      Appearance <- "PN_PB\PTMUX_F_TLN113_128"
   TextField "OBJECT_484" at 1009,421 size 40x20; Text '115'
      Appearance <- "PN_PB\PTMUX_F_TLN113_128"
   GraphicIOField "OBJECT_485" at 936,410 size 60x43; PictureList "PB_Slave_Bit12_2"
      ProcessValue <- "PN_PB\PTMUX_P_TLN113_128"
   TextField "OBJECT_486" at 946,421 size 40x20; Text '116'
      Appearance <- "PN_PB\PTMUX_F_TLN113_128"
   GraphicIOField "OBJECT_488" at 748,410 size 60x43; PictureList "PB_Slave_Bit15_2"
      ProcessValue <- "PN_PB\PTMUX_P_TLN113_128"
   TextField "OBJECT_489" at 758,421 size 40x20; Text '119'
      Appearance <- "PN_PB\PTMUX_F_TLN113_128"
   GraphicIOField "OBJECT_210" at 246,89 size 60x43; PictureList "PB_Slave_Bit7_2"
      ProcessValue <- "PN_PB\PTMUX_P_TLN1_16"
   GraphicIOField "OBJECT_214" at 372,89 size 60x43; PictureList "PB_Slave_Bit5_2"
      ProcessValue <- "PN_PB\PTMUX_P_TLN1_16"
   GraphicIOField "OBJECT_215" at 434,89 size 60x43; PictureList "PB_Slave_Bit4_2"
      ProcessValue <- "PN_PB\PTMUX_P_TLN1_16"
   TextField "OBJECT_218" at 506,100 size 40x20; Text '1'
   GraphicIOField "OBJECT_219" at 560,89 size 60x43; PictureList "PB_Slave_Bit2_2"
      ProcessValue <- "PN_PB\PTMUX_P_TLN1_16"
   GraphicIOField "OBJECT_221" at 622,89 size 60x43; PictureList "PB_Slave_Bit1_2"
      ProcessValue <- "PN_PB\PTMUX_P_TLN1_16"
   GraphicIOField "OBJECT_222" at 685,89 size 60x43; PictureList "PB_Slave_Bit0_2"
      ProcessValue <- "PN_PB\PTMUX_P_TLN1_16"
   TextField "OBJECT_223" at 696,100 size 40x20; Text '8'
      Appearance <- "PN_PB\PTMUX_F_TLN1_16"
   GraphicIOField "OBJECT_225" at 497,89 size 60x43; PictureList "PB_Slave_Bit3_2"
      ProcessValue <- "PN_PB\PTMUX_P_TLN1_16"
   TextField "OBJECT_226" at 633,100 size 40x20; Text '9'
      Appearance <- "PN_PB\PTMUX_F_TLN1_16"
   TextField "OBJECT_227" at 570,100 size 40x20; Text '10'
      Appearance <- "PN_PB\PTMUX_F_TLN1_16"
   TextField "OBJECT_228" at 508,100 size 40x20; Text '11'
      Appearance <- "PN_PB\PTMUX_F_TLN1_16"
   TextField "OBJECT_229" at 445,100 size 40x20; Text '12'
      Appearance <- "PN_PB\PTMUX_F_TLN1_16"
   TextField "OBJECT_230" at 382,100 size 40x20; Text '13'
      Appearance <- "PN_PB\PTMUX_F_TLN1_16"
   TextField "OBJECT_231" at 320,100 size 40x20; Text '14'
      Appearance <- "PN_PB\PTMUX_F_TLN1_16"
   TextField "OBJECT_232" at 257,100 size 40x20; Text '15'
      Appearance <- "PN_PB\PTMUX_F_TLN1_16"
   GraphicIOField "OBJECT_250" at 246,134 size 60x43; PictureList "PB_Slave_Bit7_2"
      ProcessValue <- "PN_PB\PTMUX_P_TLN17_32"
   GraphicIOField "OBJECT_251" at 309,134 size 60x43; PictureList "PB_Slave_Bit6_2"
      ProcessValue <- "PN_PB\PTMUX_P_TLN17_32"
   GraphicIOField "OBJECT_252" at 372,134 size 60x43; PictureList "PB_Slave_Bit5_2"
      ProcessValue <- "PN_PB\PTMUX_P_TLN17_32"
   GraphicIOField "OBJECT_253" at 434,134 size 60x43; PictureList "PB_Slave_Bit4_2"
      ProcessValue <- "PN_PB\PTMUX_P_TLN17_32"
   TextField "OBJECT_254" at 506,145 size 40x20; Text '1'
   GraphicIOField "OBJECT_255" at 560,134 size 60x43; PictureList "PB_Slave_Bit2_2"
      ProcessValue <- "PN_PB\PTMUX_P_TLN17_32"
   GraphicIOField "OBJECT_256" at 622,134 size 60x43; PictureList "PB_Slave_Bit1_2"
      ProcessValue <- "PN_PB\PTMUX_P_TLN17_32"
   GraphicIOField "OBJECT_257" at 685,134 size 60x43; PictureList "PB_Slave_Bit0_2"
      ProcessValue <- "PN_PB\PTMUX_P_TLN17_32"
   TextField "OBJECT_258" at 696,145 size 40x20; Text '24'
      Appearance <- "PN_PB\PTMUX_F_TLN17_32"
   GraphicIOField "OBJECT_259" at 497,134 size 60x43; PictureList "PB_Slave_Bit3_2"
      ProcessValue <- "PN_PB\PTMUX_P_TLN17_32"
   TextField "OBJECT_260" at 633,145 size 40x20; Text '25'
      Appearance <- "PN_PB\PTMUX_F_TLN17_32"
   TextField "OBJECT_261" at 570,145 size 40x20; Text '26'
      Appearance <- "PN_PB\PTMUX_F_TLN17_32"
   TextField "OBJECT_262" at 508,145 size 40x20; Text '27'
      Appearance <- "PN_PB\PTMUX_F_TLN17_32"
   TextField "OBJECT_263" at 445,145 size 40x20; Text '28'
      Appearance <- "PN_PB\PTMUX_F_TLN17_32"
   TextField "OBJECT_264" at 382,145 size 40x20; Text '29'
      Appearance <- "PN_PB\PTMUX_F_TLN17_32"
   TextField "OBJECT_265" at 320,145 size 40x20; Text '30'
      Appearance <- "PN_PB\PTMUX_F_TLN17_32"
   TextField "OBJECT_266" at 257,145 size 40x20; Text '31'
      Appearance <- "PN_PB\PTMUX_F_TLN17_32"
   GraphicIOField "OBJECT_283" at 246,180 size 60x43; PictureList "PB_Slave_Bit7_2"
      ProcessValue <- "PN_PB\PTMUX_P_TLN33_48"
   GraphicIOField "OBJECT_284" at 309,180 size 60x43; PictureList "PB_Slave_Bit6_2"
      ProcessValue <- "PN_PB\PTMUX_P_TLN33_48"
   GraphicIOField "OBJECT_285" at 372,180 size 60x43; PictureList "PB_Slave_Bit5_2"
      ProcessValue <- "PN_PB\PTMUX_P_TLN33_48"
   GraphicIOField "OBJECT_286" at 434,180 size 60x43; PictureList "PB_Slave_Bit4_2"
      ProcessValue <- "PN_PB\PTMUX_P_TLN33_48"
   TextField "OBJECT_287" at 506,190 size 40x20; Text '1'
   GraphicIOField "OBJECT_288" at 560,180 size 60x43; PictureList "PB_Slave_Bit2_2"
      ProcessValue <- "PN_PB\PTMUX_P_TLN33_48"
   GraphicIOField "OBJECT_289" at 622,180 size 60x43; PictureList "PB_Slave_Bit1_2"
      ProcessValue <- "PN_PB\PTMUX_P_TLN33_48"
   GraphicIOField "OBJECT_290" at 685,180 size 60x43; PictureList "PB_Slave_Bit0_2"
      ProcessValue <- "PN_PB\PTMUX_P_TLN33_48"
   TextField "OBJECT_291" at 696,190 size 40x20; Text '40'
      Appearance <- "PN_PB\PTMUX_F_TLN33_48"
   GraphicIOField "OBJECT_292" at 497,180 size 60x43; PictureList "PB_Slave_Bit3_2"
      ProcessValue <- "PN_PB\PTMUX_P_TLN33_48"
   TextField "OBJECT_293" at 633,190 size 40x20; Text '41'
      Appearance <- "PN_PB\PTMUX_F_TLN33_48"
   TextField "OBJECT_294" at 570,190 size 40x20; Text '42'
      Appearance <- "PN_PB\PTMUX_F_TLN33_48"
   TextField "OBJECT_295" at 508,190 size 40x20; Text '43'
      Appearance <- "PN_PB\PTMUX_F_TLN33_48"
   TextField "OBJECT_296" at 445,190 size 40x20; Text '44'
      Appearance <- "PN_PB\PTMUX_F_TLN33_48"
   TextField "OBJECT_297" at 382,190 size 40x20; Text '45'
      Appearance <- "PN_PB\PTMUX_F_TLN33_48"
   TextField "OBJECT_298" at 320,190 size 40x20; Text '46'
      Appearance <- "PN_PB\PTMUX_F_TLN33_48"
   TextField "OBJECT_299" at 257,190 size 40x20; Text '47'
      Appearance <- "PN_PB\PTMUX_F_TLN33_48"
   GraphicIOField "OBJECT_318" at 246,225 size 60x43; PictureList "PB_Slave_Bit7_2"
      ProcessValue <- "PN_PB\PTMUX_P_TLN49_64"
   GraphicIOField "OBJECT_319" at 309,225 size 60x43; PictureList "PB_Slave_Bit6_2"
      ProcessValue <- "PN_PB\PTMUX_P_TLN49_64"
   GraphicIOField "OBJECT_320" at 372,225 size 60x43; PictureList "PB_Slave_Bit5_2"
      ProcessValue <- "PN_PB\PTMUX_P_TLN49_64"
   GraphicIOField "OBJECT_321" at 434,225 size 60x43; PictureList "PB_Slave_Bit4_2"
      ProcessValue <- "PN_PB\PTMUX_P_TLN49_64"
   TextField "OBJECT_322" at 506,236 size 40x20; Text '1'
   GraphicIOField "OBJECT_323" at 560,225 size 60x43; PictureList "PB_Slave_Bit2_2"
      ProcessValue <- "PN_PB\PTMUX_P_TLN49_64"
   GraphicIOField "OBJECT_324" at 622,225 size 60x43; PictureList "PB_Slave_Bit1_2"
      ProcessValue <- "PN_PB\PTMUX_P_TLN49_64"
   GraphicIOField "OBJECT_325" at 685,225 size 60x43; PictureList "PB_Slave_Bit0_2"
      ProcessValue <- "PN_PB\PTMUX_P_TLN49_64"
   TextField "OBJECT_326" at 696,236 size 40x20; Text '56'
      Appearance <- "PN_PB\PTMUX_F_TLN49_64"
   GraphicIOField "OBJECT_327" at 497,225 size 60x43; PictureList "PB_Slave_Bit3_2"
      ProcessValue <- "PN_PB\PTMUX_P_TLN49_64"
   TextField "OBJECT_328" at 633,236 size 40x20; Text '57'
      Appearance <- "PN_PB\PTMUX_F_TLN49_64"
   TextField "OBJECT_329" at 570,236 size 40x20; Text '58'
      Appearance <- "PN_PB\PTMUX_F_TLN49_64"
   TextField "OBJECT_330" at 508,236 size 40x20; Text '59'
      Appearance <- "PN_PB\PTMUX_F_TLN49_64"
   TextField "OBJECT_331" at 445,236 size 40x20; Text '60'
      Appearance <- "PN_PB\PTMUX_F_TLN49_64"
   TextField "OBJECT_332" at 382,236 size 40x20; Text '61'
      Appearance <- "PN_PB\PTMUX_F_TLN49_64"
   TextField "OBJECT_333" at 320,236 size 40x20; Text '62'
      Appearance <- "PN_PB\PTMUX_F_TLN49_64"
   TextField "OBJECT_334" at 257,236 size 40x20; Text '63'
      Appearance <- "PN_PB\PTMUX_F_TLN49_64"
   GraphicIOField "OBJECT_352" at 246,270 size 60x43; PictureList "PB_Slave_Bit7_2"
      ProcessValue <- "PN_PB\PTMUX_P_TLN65_80"
   GraphicIOField "OBJECT_353" at 309,270 size 60x43; PictureList "PB_Slave_Bit6_2"
      ProcessValue <- "PN_PB\PTMUX_P_TLN65_80"
   GraphicIOField "OBJECT_354" at 372,270 size 60x43; PictureList "PB_Slave_Bit5_2"
      ProcessValue <- "PN_PB\PTMUX_P_TLN65_80"
   GraphicIOField "OBJECT_355" at 434,270 size 60x43; PictureList "PB_Slave_Bit4_2"
      ProcessValue <- "PN_PB\PTMUX_P_TLN65_80"
   TextField "OBJECT_356" at 506,282 size 40x20; Text '1'
   GraphicIOField "OBJECT_357" at 560,270 size 60x43; PictureList "PB_Slave_Bit2_2"
      ProcessValue <- "PN_PB\PTMUX_P_TLN65_80"
   GraphicIOField "OBJECT_358" at 622,270 size 60x43; PictureList "PB_Slave_Bit1_2"
      ProcessValue <- "PN_PB\PTMUX_P_TLN65_80"
   GraphicIOField "OBJECT_359" at 685,270 size 60x43; PictureList "PB_Slave_Bit0_2"
      ProcessValue <- "PN_PB\PTMUX_P_TLN65_80"
   TextField "OBJECT_360" at 696,282 size 40x20; Text '72'
      Appearance <- "PN_PB\PTMUX_F_TLN65_80"
   GraphicIOField "OBJECT_361" at 497,270 size 60x43; PictureList "PB_Slave_Bit3_2"
      ProcessValue <- "PN_PB\PTMUX_P_TLN65_80"
   TextField "OBJECT_362" at 633,282 size 40x20; Text '73'
      Appearance <- "PN_PB\PTMUX_F_TLN65_80"
   TextField "OBJECT_363" at 570,282 size 40x20; Text '74'
      Appearance <- "PN_PB\PTMUX_F_TLN65_80"
   TextField "OBJECT_364" at 508,282 size 40x20; Text '75'
      Appearance <- "PN_PB\PTMUX_F_TLN65_80"
   TextField "OBJECT_365" at 445,282 size 40x20; Text '76'
      Appearance <- "PN_PB\PTMUX_F_TLN65_80"
   TextField "OBJECT_366" at 382,282 size 40x20; Text '77'
      Appearance <- "PN_PB\PTMUX_F_TLN65_80"
   TextField "OBJECT_367" at 320,282 size 40x20; Text '78'
      Appearance <- "PN_PB\PTMUX_F_TLN65_80"
   TextField "OBJECT_368" at 257,282 size 40x20; Text '79'
      Appearance <- "PN_PB\PTMUX_F_TLN65_80"
   GraphicIOField "OBJECT_388" at 246,317 size 60x43; PictureList "PB_Slave_Bit7_2"
      ProcessValue <- "PN_PB\PTMUX_P_TLN81_96"
   GraphicIOField "OBJECT_389" at 309,317 size 60x43; PictureList "PB_Slave_Bit6_2"
      ProcessValue <- "PN_PB\PTMUX_P_TLN81_96"
   GraphicIOField "OBJECT_390" at 372,317 size 60x43; PictureList "PB_Slave_Bit5_2"
      ProcessValue <- "PN_PB\PTMUX_P_TLN81_96"
   GraphicIOField "OBJECT_391" at 434,317 size 60x43; PictureList "PB_Slave_Bit4_2"
      ProcessValue <- "PN_PB\PTMUX_P_TLN81_96"
   TextField "OBJECT_392" at 506,329 size 40x20; Text '1'
   GraphicIOField "OBJECT_393" at 560,317 size 60x43; PictureList "PB_Slave_Bit2_2"
      ProcessValue <- "PN_PB\PTMUX_P_TLN81_96"
   GraphicIOField "OBJECT_394" at 622,317 size 60x43; PictureList "PB_Slave_Bit1_2"
      ProcessValue <- "PN_PB\PTMUX_P_TLN81_96"
   GraphicIOField "OBJECT_395" at 685,317 size 60x43; PictureList "PB_Slave_Bit0_2"
      ProcessValue <- "PN_PB\PTMUX_P_TLN81_96"
   TextField "OBJECT_396" at 696,329 size 40x20; Text '88'
      Appearance <- "PN_PB\PTMUX_F_TLN81_96"
   GraphicIOField "OBJECT_397" at 497,317 size 60x43; PictureList "PB_Slave_Bit3_2"
      ProcessValue <- "PN_PB\PTMUX_P_TLN81_96"
   TextField "OBJECT_398" at 633,329 size 40x20; Text '89'
      Appearance <- "PN_PB\PTMUX_F_TLN81_96"
   TextField "OBJECT_399" at 570,329 size 40x20; Text '90'
      Appearance <- "PN_PB\PTMUX_F_TLN81_96"
   TextField "OBJECT_400" at 508,329 size 40x20; Text '91'
      Appearance <- "PN_PB\PTMUX_F_TLN81_96"
   TextField "OBJECT_401" at 445,329 size 40x20; Text '92'
      Appearance <- "PN_PB\PTMUX_F_TLN81_96"
   TextField "OBJECT_402" at 382,329 size 40x20; Text '93'
      Appearance <- "PN_PB\PTMUX_F_TLN81_96"
   TextField "OBJECT_403" at 320,329 size 40x20; Text '94'
      Appearance <- "PN_PB\PTMUX_F_TLN81_96"
   TextField "OBJECT_404" at 257,329 size 40x20; Text '95'
      Appearance <- "PN_PB\PTMUX_F_TLN81_96"
   GraphicIOField "OBJECT_423" at 246,364 size 60x43; PictureList "PB_Slave_Bit7_2"
      ProcessValue <- "PN_PB\PTMUX_P_TLN97_112"
   GraphicIOField "OBJECT_424" at 309,364 size 60x43; PictureList "PB_Slave_Bit6_2"
      ProcessValue <- "PN_PB\PTMUX_P_TLN97_112"
   GraphicIOField "OBJECT_425" at 372,364 size 60x43; PictureList "PB_Slave_Bit5_2"
      ProcessValue <- "PN_PB\PTMUX_P_TLN97_112"
   GraphicIOField "OBJECT_426" at 434,364 size 60x43; PictureList "PB_Slave_Bit4_2"
      ProcessValue <- "PN_PB\PTMUX_P_TLN97_112"
   TextField "OBJECT_427" at 506,376 size 40x20; Text '1'
   GraphicIOField "OBJECT_428" at 560,364 size 60x43; PictureList "PB_Slave_Bit2_2"
      ProcessValue <- "PN_PB\PTMUX_P_TLN97_112"
   GraphicIOField "OBJECT_429" at 622,364 size 60x43; PictureList "PB_Slave_Bit1_2"
      ProcessValue <- "PN_PB\PTMUX_P_TLN97_112"
   GraphicIOField "OBJECT_430" at 685,364 size 60x43; PictureList "PB_Slave_Bit0_2"
      ProcessValue <- "PN_PB\PTMUX_P_TLN97_112"
   TextField "OBJECT_431" at 696,376 size 40x20; Text '104'
      Appearance <- "PN_PB\PTMUX_F_TLN97_112"
   GraphicIOField "OBJECT_432" at 497,364 size 60x43; PictureList "PB_Slave_Bit3_2"
      ProcessValue <- "PN_PB\PTMUX_P_TLN97_112"
   TextField "OBJECT_433" at 633,376 size 40x20; Text '105'
      Appearance <- "PN_PB\PTMUX_F_TLN97_112"
   TextField "OBJECT_434" at 570,376 size 40x20; Text '106'
      Appearance <- "PN_PB\PTMUX_F_TLN97_112"
   TextField "OBJECT_435" at 508,376 size 40x20; Text '107'
      Appearance <- "PN_PB\PTMUX_F_TLN97_112"
   TextField "OBJECT_436" at 445,376 size 40x20; Text '108'
      Appearance <- "PN_PB\PTMUX_F_TLN97_112"
   TextField "OBJECT_437" at 382,376 size 40x20; Text '109'
      Appearance <- "PN_PB\PTMUX_F_TLN97_112"
   TextField "OBJECT_438" at 320,376 size 40x20; Text '110'
      Appearance <- "PN_PB\PTMUX_F_TLN97_112"
   TextField "OBJECT_439" at 257,376 size 40x20; Text '111'
      Appearance <- "PN_PB\PTMUX_F_TLN97_112"
   GraphicIOField "OBJECT_460" at 309,410 size 60x43; PictureList "PB_Slave_Bit6_2"
      ProcessValue <- "PN_PB\PTMUX_P_TLN113_128"
   GraphicIOField "OBJECT_461" at 372,410 size 60x43; PictureList "PB_Slave_Bit5_2"
      ProcessValue <- "PN_PB\PTMUX_P_TLN113_128"
   GraphicIOField "OBJECT_462" at 434,410 size 60x43; PictureList "PB_Slave_Bit4_2"
      ProcessValue <- "PN_PB\PTMUX_P_TLN113_128"
   TextField "OBJECT_463" at 506,421 size 40x20; Text '1'
   GraphicIOField "OBJECT_464" at 559,410 size 60x43; PictureList "PB_Slave_Bit2_2"
      ProcessValue <- "PN_PB\PTMUX_P_TLN113_128"
   GraphicIOField "OBJECT_465" at 622,410 size 60x43; PictureList "PB_Slave_Bit1_2"
      ProcessValue <- "PN_PB\PTMUX_P_TLN113_128"
   GraphicIOField "OBJECT_466" at 685,410 size 60x43; PictureList "PB_Slave_Bit0_2"
      ProcessValue <- "PN_PB\PTMUX_P_TLN113_128"
   TextField "OBJECT_467" at 696,421 size 40x20; Text '120'
      Appearance <- "PN_PB\PTMUX_F_TLN113_128"
   GraphicIOField "OBJECT_468" at 497,410 size 60x43; PictureList "PB_Slave_Bit3_2"
      ProcessValue <- "PN_PB\PTMUX_P_TLN113_128"
   TextField "OBJECT_469" at 633,421 size 40x20; Text '121'
      Appearance <- "PN_PB\PTMUX_F_TLN113_128"
   TextField "OBJECT_470" at 570,421 size 40x20; Text '122'
      Appearance <- "PN_PB\PTMUX_F_TLN113_128"
   TextField "OBJECT_471" at 508,421 size 40x20; Text '123'
      Appearance <- "PN_PB\PTMUX_F_TLN113_128"
   TextField "OBJECT_472" at 445,421 size 40x20; Text '124'
      Appearance <- "PN_PB\PTMUX_F_TLN113_128"
   TextField "OBJECT_473" at 382,421 size 40x20; Text '125'
      Appearance <- "PN_PB\PTMUX_F_TLN113_128"
   TextField "OBJECT_474" at 320,421 size 40x20; Text '126'
      Appearance <- "PN_PB\PTMUX_F_TLN113_128"
   GraphicIOField "OBJECT_490" at 246,410 size 60x43; PictureList "PB_Slave_Bit7_2"
      ProcessValue <- "PN_PB\PTMUX_P_TLN113_128"
   TextField "OBJECT_491" at 257,421 size 40x20; Text '127'
      Appearance <- "PN_PB\PTMUX_F_TLN113_128"
   TextField "OBJECT_670" at 919,469 size 111x35; Text 'Legende:'
   IOField "OBJECT_111" at 524,45 size 47x29; FormatPattern 999
      ProcessValue <- "PN_PB\IO_Sys_ID"
   GraphicIOField "OBJECT_5" at 873,89 size 60x43; PictureList "PB_Slave_Bit13_2"
      ProcessValue <- "PN_PB\PTMUX_P_TLN1_16"
   TextField "OBJECT_238" at 884,100 size 40x20; Text '5'
      Appearance <- "PN_PB\PTMUX_F_TLN1_16"
   TextField "OBJECT_513" at 255,505 size 104x29; Text 'Ort:'
   TextField "OBJECT_514" at 255,535 size 104x31; Text 'Typ:'
   TextField "OBJECT_515" at 255,565 size 131x29; Text 'Bezeichnung:'
   IOField "OBJECT_516" at 399,505 size 167x29; FormatPattern ????????????
      ProcessValue <- "PN_PB\Teiln_Nr_Ort"
   IOField "OBJECT_517" at 399,535 size 156x31; FormatPattern ????????????
      ProcessValue <- "PN_PB\Teiln_Nr_Typ"
   IOField "OBJECT_518" at 399,565 size 253x29; FormatPattern ????????????????????
      ProcessValue <- "PN_PB\Teiln_Nr_Bez"
   IOField "OBJECT_658" at 483,475 size 57x27; FormatPattern 999
      ProcessValue <- "PN_PB\PN\Teiln_Nr"
      Appearance <- "Trigger"
   TextField "OBJECT_679" at 587,475 size 67x25; Text 'Trigger'
      Appearance <- "Trigger"
   Group "Group" at 248,181 size 999x45
   Group "Group_1" at 246,92 size 999x40
   Group "Group_2" at 246,135 size 999x40
   Group "Group_3" at 246,226 size 999x40
   Group "Group_4" at 247,272 size 999x40
   Group "Group_5" at 248,319 size 999x40
   Group "Group_6" at 248,366 size 999x40
   Group "Group_7" at 248,412 size 999x40
   Button "Schaltfläche_4" at 1187,181 size 60x40; TextOff 'Text'
      on Click: SetTag("PN_PB\PN\Teiln_Nr", 32)
   Button "Schaltfläche_5" at 1126,181 size 60x40; TextOff 'Text'
      on Click: SetTag("PN_PB\PN\Teiln_Nr", 33)
   Button "Schaltfläche_6" at 1064,181 size 60x40; TextOff 'Text'
      on Click: SetTag("PN_PB\PN\Teiln_Nr", 34)
   Button "Schaltfläche_7" at 1001,181 size 60x40; TextOff 'Text'
      on Click: SetTag("PN_PB\PN\Teiln_Nr", 35)
   Button "Schaltfläche_8" at 939,181 size 60x40; TextOff 'Text'
      on Click: SetTag("PN_PB\PN\Teiln_Nr", 36)
   Button "Schaltfläche_9" at 875,181 size 60x40; TextOff 'Text'
      on Click: SetTag("PN_PB\PN\Teiln_Nr", 37)
   Button "Schaltfläche_10" at 812,181 size 60x40; TextOff 'Text'
      on Click: SetTag("PN_PB\PN\Teiln_Nr", 38)
   Button "Schaltfläche_11" at 746,186 size 60x40; TextOff 'Text'
      on Click: SetTag("PN_PB\PN\Teiln_Nr", 39)
   Button "Schaltfläche_13" at 687,181 size 60x40; TextOff 'Text'
      on Click: SetTag("PN_PB\PN\Teiln_Nr", 40)
   Button "Schaltfläche_14" at 624,181 size 60x40; TextOff 'Text'
      on Click: SetTag("PN_PB\PN\Teiln_Nr", 41)
   Button "Schaltfläche_15" at 562,181 size 60x40; TextOff 'Text'
      on Click: SetTag("PN_PB\PN\Teiln_Nr", 42)
   Button "Schaltfläche_16" at 499,181 size 60x40; TextOff 'Text'
      on Click: SetTag("PN_PB\PN\Teiln_Nr", 43)
   Button "Schaltfläche_17" at 436,181 size 60x40; TextOff 'Text'
      on Click: SetTag("PN_PB\PN\Teiln_Nr", 44)
   Button "Schaltfläche_18" at 374,181 size 60x40; TextOff 'Text'
      on Click: SetTag("PN_PB\PN\Teiln_Nr", 45)
   Button "Schaltfläche_19" at 312,181 size 60x40; TextOff 'Text'
      on Click: SetTag("PN_PB\PN\Teiln_Nr", 46)
   Button "Schaltfläche_20" at 248,181 size 60x40; TextOff 'Text'
      on Click: SetTag("PN_PB\PN\Teiln_Nr", 47)
   Button "Schaltfläche_21" at 1185,92 size 60x40; TextOff 'Text'
      on Click: SetTag("PN_PB\PN\Teiln_Nr", 0)
   Button "Schaltfläche_22" at 1124,92 size 60x40; TextOff 'Text'
      on Click: SetTag("PN_PB\PN\Teiln_Nr", 1)
   Button "Schaltfläche_23" at 1062,92 size 60x40; TextOff 'Text'
      on Click: SetTag("PN_PB\PN\Teiln_Nr", 2)
   Button "Schaltfläche_24" at 999,92 size 60x40; TextOff 'Text'
      on Click: SetTag("PN_PB\PN\Teiln_Nr", 3)
   Button "Schaltfläche_25" at 937,92 size 60x40; TextOff 'Text'
      on Click: SetTag("PN_PB\PN\Teiln_Nr", 4)
   Button "Schaltfläche_26" at 873,92 size 60x40; TextOff 'Text'
      on Click: SetTag("PN_PB\PN\Teiln_Nr", 5)
   Button "Schaltfläche_27" at 810,92 size 60x40; TextOff 'Text'
      on Click: SetTag("PN_PB\PN\Teiln_Nr", 6)
   Button "Schaltfläche_28" at 748,92 size 60x40; TextOff 'Text'
      on Click: SetTag("PN_PB\PN\Teiln_Nr", 7)
   Button "Schaltfläche_29" at 685,92 size 60x40; TextOff 'Text'
      on Click: SetTag("PN_PB\PN\Teiln_Nr", 8)
   Button "Schaltfläche_30" at 622,92 size 60x40; TextOff 'Text'
      on Click: SetTag("PN_PB\PN\Teiln_Nr", 9)
   Button "Schaltfläche_31" at 560,92 size 60x40; TextOff 'Text'
      on Click: SetTag("PN_PB\PN\Teiln_Nr", 10)
   Button "Schaltfläche_32" at 497,92 size 60x40; TextOff 'Text'
      on Click: SetTag("PN_PB\PN\Teiln_Nr", 11)
   Button "Schaltfläche_33" at 434,92 size 60x40; TextOff 'Text'
      on Click: SetTag("PN_PB\PN\Teiln_Nr", 12)
   Button "Schaltfläche_34" at 372,92 size 60x40; TextOff 'Text'
      on Click: SetTag("PN_PB\PN\Teiln_Nr", 13)
   Button "Schaltfläche_35" at 310,92 size 60x40; TextOff 'Text'
      on Click: SetTag("PN_PB\PN\Teiln_Nr", 14)
   Button "Schaltfläche_36" at 246,92 size 60x40; TextOff 'Text'
      on Click: SetTag("PN_PB\PN\Teiln_Nr", 15)
   Button "Schaltfläche_12" at 1185,135 size 60x40; TextOff 'Text'
      on Click: SetTag("PN_PB\PN\Teiln_Nr", 16)
   Button "Schaltfläche_37" at 1124,135 size 60x40; TextOff 'Text'
      on Click: SetTag("PN_PB\PN\Teiln_Nr", 17)
   Button "Schaltfläche_38" at 1062,135 size 60x40; TextOff 'Text'
      on Click: SetTag("PN_PB\PN\Teiln_Nr", 18)
   Button "Schaltfläche_39" at 999,135 size 60x40; TextOff 'Text'
      on Click: SetTag("PN_PB\PN\Teiln_Nr", 19)
   Button "Schaltfläche_40" at 937,135 size 60x40; TextOff 'Text'
      on Click: SetTag("PN_PB\PN\Teiln_Nr", 20)
   Button "Schaltfläche_41" at 873,135 size 60x40; TextOff 'Text'
      on Click: SetTag("PN_PB\PN\Teiln_Nr", 21)
   Button "Schaltfläche_42" at 810,135 size 60x40; TextOff 'Text'
      on Click: SetTag("PN_PB\PN\Teiln_Nr", 22)
   Button "Schaltfläche_43" at 748,135 size 60x40; TextOff 'Text'
      on Click: SetTag("PN_PB\PN\Teiln_Nr", 23)
   Button "Schaltfläche_44" at 685,135 size 60x40; TextOff 'Text'
      on Click: SetTag("PN_PB\PN\Teiln_Nr", 24)
   Button "Schaltfläche_45" at 622,135 size 60x40; TextOff 'Text'
      on Click: SetTag("PN_PB\PN\Teiln_Nr", 25)
   Button "Schaltfläche_46" at 560,135 size 60x40; TextOff 'Text'
      on Click: SetTag("PN_PB\PN\Teiln_Nr", 26)
   Button "Schaltfläche_47" at 497,135 size 60x40; TextOff 'Text'
      on Click: SetTag("PN_PB\PN\Teiln_Nr", 27)
   Button "Schaltfläche_48" at 434,135 size 60x40; TextOff 'Text'
      on Click: SetTag("PN_PB\PN\Teiln_Nr", 28)
   Button "Schaltfläche_49" at 372,135 size 60x40; TextOff 'Text'
      on Click: SetTag("PN_PB\PN\Teiln_Nr", 29)
   Button "Schaltfläche_50" at 310,135 size 60x40; TextOff 'Text'
      on Click: SetTag("PN_PB\PN\Teiln_Nr", 30)
   Button "Schaltfläche_51" at 246,135 size 60x40; TextOff 'Text'
      on Click: SetTag("PN_PB\PN\Teiln_Nr", 31)
   Button "Schaltfläche_52" at 1185,226 size 60x40; TextOff 'Text'
      on Click: SetTag("PN_PB\PN\Teiln_Nr", 48)
   Button "Schaltfläche_53" at 1124,226 size 60x40; TextOff 'Text'
      on Click: SetTag("PN_PB\PN\Teiln_Nr", 49)
   Button "Schaltfläche_54" at 1062,226 size 60x40; TextOff 'Text'
      on Click: SetTag("PN_PB\PN\Teiln_Nr", 50)
   Button "Schaltfläche_55" at 999,226 size 60x40; TextOff 'Text'
      on Click: SetTag("PN_PB\PN\Teiln_Nr", 51)
   Button "Schaltfläche_56" at 937,226 size 60x40; TextOff 'Text'
      on Click: SetTag("PN_PB\PN\Teiln_Nr", 52)
   Button "Schaltfläche_57" at 873,226 size 60x40; TextOff 'Text'
      on Click: SetTag("PN_PB\PN\Teiln_Nr", 53)
   Button "Schaltfläche_58" at 810,226 size 60x40; TextOff 'Text'
      on Click: SetTag("PN_PB\PN\Teiln_Nr", 54)
   Button "Schaltfläche_59" at 748,226 size 60x40; TextOff 'Text'
      on Click: SetTag("PN_PB\PN\Teiln_Nr", 55)
   Button "Schaltfläche_60" at 685,226 size 60x40; TextOff 'Text'
      on Click: SetTag("PN_PB\PN\Teiln_Nr", 56)
   Button "Schaltfläche_61" at 622,226 size 60x40; TextOff 'Text'
      on Click: SetTag("PN_PB\PN\Teiln_Nr", 57)
   Button "Schaltfläche_62" at 560,226 size 60x40; TextOff 'Text'
      on Click: SetTag("PN_PB\PN\Teiln_Nr", 58)
   Button "Schaltfläche_63" at 497,226 size 60x40; TextOff 'Text'
      on Click: SetTag("PN_PB\PN\Teiln_Nr", 59)
   Button "Schaltfläche_64" at 434,226 size 60x40; TextOff 'Text'
      on Click: SetTag("PN_PB\PN\Teiln_Nr", 60)
   Button "Schaltfläche_65" at 372,226 size 60x40; TextOff 'Text'
      on Click: SetTag("PN_PB\PN\Teiln_Nr", 61)
   Button "Schaltfläche_66" at 310,226 size 60x40; TextOff 'Text'
      on Click: SetTag("PN_PB\PN\Teiln_Nr", 62)
   Button "Schaltfläche_67" at 246,226 size 60x40; TextOff 'Text'
      on Click: SetTag("PN_PB\PN\Teiln_Nr", 63)
   Button "Schaltfläche_68" at 1186,272 size 60x40; TextOff 'Text'
      on Click: SetTag("PN_PB\PN\Teiln_Nr", 64)
   Button "Schaltfläche_69" at 1125,272 size 60x40; TextOff 'Text'
      on Click: SetTag("PN_PB\PN\Teiln_Nr", 65)
   Button "Schaltfläche_70" at 1063,272 size 60x40; TextOff 'Text'
      on Click: SetTag("PN_PB\PN\Teiln_Nr", 66)
   Button "Schaltfläche_71" at 1000,272 size 60x40; TextOff 'Text'
      on Click: SetTag("PN_PB\PN\Teiln_Nr", 67)
   Button "Schaltfläche_72" at 938,272 size 60x40; TextOff 'Text'
      on Click: SetTag("PN_PB\PN\Teiln_Nr", 68)
   Button "Schaltfläche_73" at 874,272 size 60x40; TextOff 'Text'
      on Click: SetTag("PN_PB\PN\Teiln_Nr", 69)
   Button "Schaltfläche_74" at 811,272 size 60x40; TextOff 'Text'
      on Click: SetTag("PN_PB\PN\Teiln_Nr", 70)
   Button "Schaltfläche_75" at 749,272 size 60x40; TextOff 'Text'
      on Click: SetTag("PN_PB\PN\Teiln_Nr", 71)
   Button "Schaltfläche_76" at 686,272 size 60x40; TextOff 'Text'
      on Click: SetTag("PN_PB\PN\Teiln_Nr", 72)
   Button "Schaltfläche_77" at 623,272 size 60x40; TextOff 'Text'
      on Click: SetTag("PN_PB\PN\Teiln_Nr", 73)
   Button "Schaltfläche_78" at 561,272 size 60x40; TextOff 'Text'
      on Click: SetTag("PN_PB\PN\Teiln_Nr", 74)
   Button "Schaltfläche_79" at 498,272 size 60x40; TextOff 'Text'
      on Click: SetTag("PN_PB\PN\Teiln_Nr", 75)
   Button "Schaltfläche_80" at 435,272 size 60x40; TextOff 'Text'
      on Click: SetTag("PN_PB\PN\Teiln_Nr", 76)
   Button "Schaltfläche_81" at 373,272 size 60x40; TextOff 'Text'
      on Click: SetTag("PN_PB\PN\Teiln_Nr", 77)
   Button "Schaltfläche_82" at 311,272 size 60x40; TextOff 'Text'
      on Click: SetTag("PN_PB\PN\Teiln_Nr", 78)
   Button "Schaltfläche_83" at 247,272 size 60x40; TextOff 'Text'
      on Click: SetTag("PN_PB\PN\Teiln_Nr", 79)
   Button "Schaltfläche_84" at 1187,319 size 60x40; TextOff 'Text'
      on Click: SetTag("PN_PB\PN\Teiln_Nr", 80)
   Button "Schaltfläche_85" at 1126,319 size 60x40; TextOff 'Text'
      on Click: SetTag("PN_PB\PN\Teiln_Nr", 81)
   Button "Schaltfläche_86" at 1064,319 size 60x40; TextOff 'Text'
      on Click: SetTag("PN_PB\PN\Teiln_Nr", 82)
   Button "Schaltfläche_87" at 1001,319 size 60x40; TextOff 'Text'
      on Click: SetTag("PN_PB\PN\Teiln_Nr", 83)
   Button "Schaltfläche_88" at 939,319 size 60x40; TextOff 'Text'
      on Click: SetTag("PN_PB\PN\Teiln_Nr", 84)
   Button "Schaltfläche_89" at 875,319 size 60x40; TextOff 'Text'
      on Click: SetTag("PN_PB\PN\Teiln_Nr", 85)
   Button "Schaltfläche_90" at 812,319 size 60x40; TextOff 'Text'
      on Click: SetTag("PN_PB\PN\Teiln_Nr", 86)
   Button "Schaltfläche_91" at 750,319 size 60x40; TextOff 'Text'
      on Click: SetTag("PN_PB\PN\Teiln_Nr", 87)
   Button "Schaltfläche_92" at 687,319 size 60x40; TextOff 'Text'
      on Click: SetTag("PN_PB\PN\Teiln_Nr", 88)
   Button "Schaltfläche_93" at 624,319 size 60x40; TextOff 'Text'
      on Click: SetTag("PN_PB\PN\Teiln_Nr", 89)
   Button "Schaltfläche_94" at 562,319 size 60x40; TextOff 'Text'
      on Click: SetTag("PN_PB\PN\Teiln_Nr", 90)
   Button "Schaltfläche_95" at 499,319 size 60x40; TextOff 'Text'
      on Click: SetTag("PN_PB\PN\Teiln_Nr", 91)
   Button "Schaltfläche_96" at 436,319 size 60x40; TextOff 'Text'
      on Click: SetTag("PN_PB\PN\Teiln_Nr", 92)
   Button "Schaltfläche_97" at 374,319 size 60x40; TextOff 'Text'
      on Click: SetTag("PN_PB\PN\Teiln_Nr", 93)
   Button "Schaltfläche_98" at 312,319 size 60x40; TextOff 'Text'
      on Click: SetTag("PN_PB\PN\Teiln_Nr", 94)
   Button "Schaltfläche_99" at 248,319 size 60x40; TextOff 'Text'
      on Click: SetTag("PN_PB\PN\Teiln_Nr", 95)
   Button "Schaltfläche_100" at 1187,366 size 60x40; TextOff 'Text'
      on Click: SetTag("PN_PB\PN\Teiln_Nr", 96)
   Button "Schaltfläche_101" at 1126,366 size 60x40; TextOff 'Text'
      on Click: SetTag("PN_PB\PN\Teiln_Nr", 97)
   Button "Schaltfläche_102" at 1064,366 size 60x40; TextOff 'Text'
      on Click: SetTag("PN_PB\PN\Teiln_Nr", 98)
   Button "Schaltfläche_103" at 1001,366 size 60x40; TextOff 'Text'
      on Click: SetTag("PN_PB\PN\Teiln_Nr", 99)
   Button "Schaltfläche_104" at 939,366 size 60x40; TextOff 'Text'
      on Click: SetTag("PN_PB\PN\Teiln_Nr", 100)
   Button "Schaltfläche_105" at 875,366 size 60x40; TextOff 'Text'
      on Click: SetTag("PN_PB\PN\Teiln_Nr", 101)
   Button "Schaltfläche_106" at 812,366 size 60x40; TextOff 'Text'
      on Click: SetTag("PN_PB\PN\Teiln_Nr", 102)
   Button "Schaltfläche_107" at 750,366 size 60x40; TextOff 'Text'
      on Click: SetTag("PN_PB\PN\Teiln_Nr", 103)
   Button "Schaltfläche_108" at 687,366 size 60x40; TextOff 'Text'
      on Click: SetTag("PN_PB\PN\Teiln_Nr", 104)
   Button "Schaltfläche_109" at 624,366 size 60x40; TextOff 'Text'
      on Click: SetTag("PN_PB\PN\Teiln_Nr", 105)
   Button "Schaltfläche_110" at 562,366 size 60x40; TextOff 'Text'
      on Click: SetTag("PN_PB\PN\Teiln_Nr", 106)
   Button "Schaltfläche_111" at 499,366 size 60x40; TextOff 'Text'
      on Click: SetTag("PN_PB\PN\Teiln_Nr", 107)
   Button "Schaltfläche_112" at 436,366 size 60x40; TextOff 'Text'
      on Click: SetTag("PN_PB\PN\Teiln_Nr", 108)
   Button "Schaltfläche_113" at 374,366 size 60x40; TextOff 'Text'
      on Click: SetTag("PN_PB\PN\Teiln_Nr", 109)
   Button "Schaltfläche_114" at 312,366 size 60x40; TextOff 'Text'
      on Click: SetTag("PN_PB\PN\Teiln_Nr", 110)
   Button "Schaltfläche_115" at 248,366 size 60x40; TextOff 'Text'
      on Click: SetTag("PN_PB\PN\Teiln_Nr", 111)
   Button "Schaltfläche_116" at 1187,412 size 60x40; TextOff 'Text'
      on Click: SetTag("PN_PB\PN\Teiln_Nr", 112)
   Button "Schaltfläche_117" at 1126,412 size 60x40; TextOff 'Text'
      on Click: SetTag("PN_PB\PN\Teiln_Nr", 113)
   Button "Schaltfläche_118" at 1064,412 size 60x40; TextOff 'Text'
      on Click: SetTag("PN_PB\PN\Teiln_Nr", 114)
   Button "Schaltfläche_119" at 1001,412 size 60x40; TextOff 'Text'
      on Click: SetTag("PN_PB\PN\Teiln_Nr", 115)
   Button "Schaltfläche_120" at 939,412 size 60x40; TextOff 'Text'
      on Click: SetTag("PN_PB\PN\Teiln_Nr", 116)
   Button "Schaltfläche_121" at 875,412 size 60x40; TextOff 'Text'
      on Click: SetTag("PN_PB\PN\Teiln_Nr", 117)
   Button "Schaltfläche_122" at 812,412 size 60x40; TextOff 'Text'
      on Click: SetTag("PN_PB\PN\Teiln_Nr", 118)
   Button "Schaltfläche_123" at 750,412 size 60x40; TextOff 'Text'
      on Click: SetTag("PN_PB\PN\Teiln_Nr", 119)
   Button "Schaltfläche_124" at 687,412 size 60x40; TextOff 'Text'
      on Click: SetTag("PN_PB\PN\Teiln_Nr", 120)
   Button "Schaltfläche_125" at 624,412 size 60x40; TextOff 'Text'
      on Click: SetTag("PN_PB\PN\Teiln_Nr", 121)
   Button "Schaltfläche_126" at 562,412 size 60x40; TextOff 'Text'
      on Click: SetTag("PN_PB\PN\Teiln_Nr", 122)
   Button "Schaltfläche_127" at 499,412 size 60x40; TextOff 'Text'
      on Click: SetTag("PN_PB\PN\Teiln_Nr", 123)
   Button "Schaltfläche_128" at 436,412 size 60x40; TextOff 'Text'
      on Click: SetTag("PN_PB\PN\Teiln_Nr", 124)
   Button "Schaltfläche_129" at 374,412 size 60x40; TextOff 'Text'
      on Click: SetTag("PN_PB\PN\Teiln_Nr", 125)
   Button "Schaltfläche_130" at 312,412 size 60x40; TextOff 'Text'
      on Click: SetTag("PN_PB\PN\Teiln_Nr", 126)
   Button "Schaltfläche_131" at 248,412 size 60x40; TextOff 'Text'
      on Click: SetTag("PN_PB\PN\Teiln_Nr", 127)

